REGION Network 151: PRODUCTION HOLD PB NOT RESET
   RUNG wire#powerrail
      Contact( "reset" )
      { S7_Templates := "SrcType := Word" } EQ_Contact(in1 := "DB101_DB_SDC_FAULTS".Carrier_Fault[44], in2 := 103)
      Coil( "DB302_HMI_Faults".Carrier44_Faults_3.%X14 )
   END_RUNG
   // the same network as SCL:
   "DB302_HMI_Faults".Carrier44_Faults_3.%X14 := "reset" AND ("DB101_DB_SDC_FAULTS".Carrier_Fault[44] = 103);
END_REGION

REGION Network 152: CARRIER FAULTS MASKED
   Label( C44_Comm_Flt )
   RUNG wire#powerrail
      Contact( "EMS".Carrier[44].FaultsMasked )
      Coil( "DB302_HMI_Faults".Carrier44_Faults_3.%X15 )
   END_RUNG
   // the same network as SCL:
   C44_Comm_Flt:
   "DB302_HMI_Faults".Carrier44_Faults_3.%X15 := "EMS".Carrier[44].FaultsMasked;
END_REGION

REGION Network 153: CARRIER 45 FAULTS
END_REGION

REGION Network 154: CARRIER PLC NOT COMMUNICATING
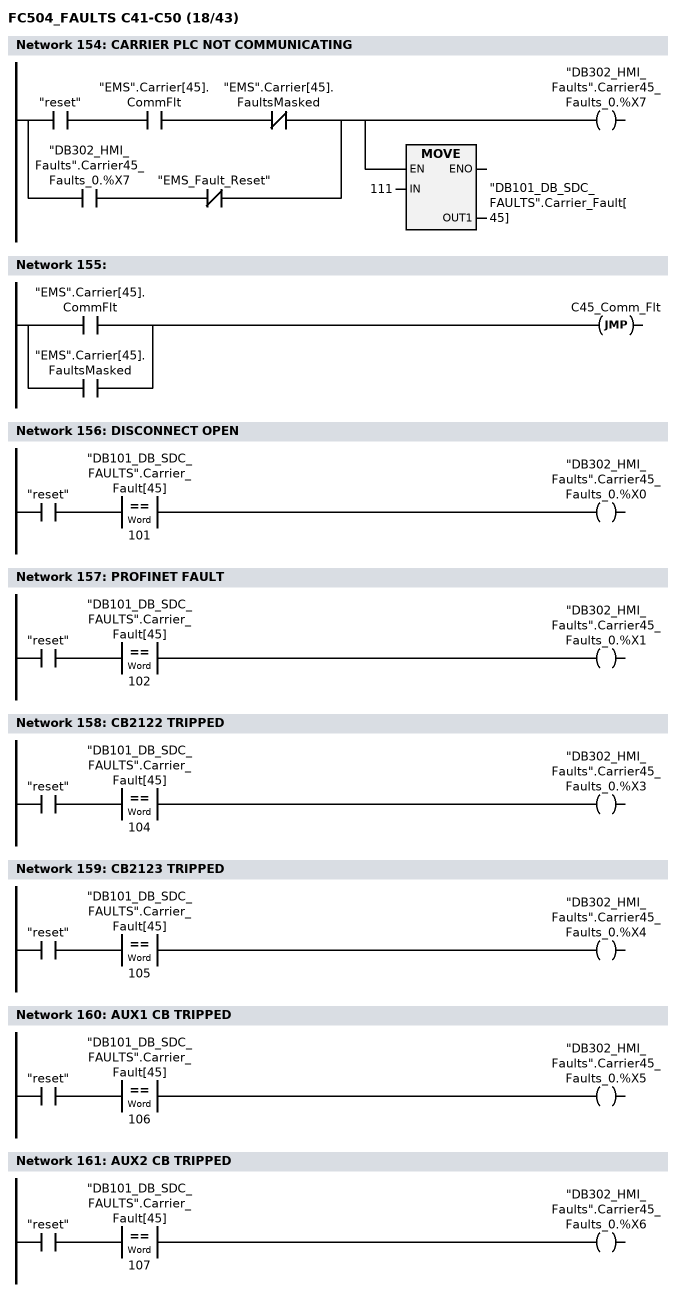
   RUNG wire#powerrail
      Contact( "reset" )
      Contact( "EMS".Carrier[45].CommFlt )
      I_Contact( "EMS".Carrier[45].FaultsMasked )
      wire#w1
      Coil( "DB302_HMI_Faults".Carrier45_Faults_0.%X7 )
   END_RUNG
   RUNG wire#powerrail
      Contact( "DB302_HMI_Faults".Carrier45_Faults_0.%X7 )
      I_Contact( "EMS_Fault_Reset" )
   END_RUNG wire#w1
   RUNG wire#w1
      Move(in := 111, out1 => "DB101_DB_SDC_FAULTS".Carrier_Fault[45])
   END_RUNG
   // the same network as SCL:
   "DB302_HMI_Faults".Carrier45_Faults_0.%X7 := ("reset" AND "EMS".Carrier[45].CommFlt AND NOT "EMS".Carrier[45].FaultsMasked) OR ("DB302_HMI_Faults".Carrier45_Faults_0.%X7 AND NOT "EMS_Fault_Reset");
   IF "DB302_HMI_Faults".Carrier45_Faults_0.%X7 THEN "DB101_DB_SDC_FAULTS".Carrier_Fault[45] := 111; END_IF;
END_REGION

REGION Network 155
   RUNG wire#powerrail
      Contact( "EMS".Carrier[45].CommFlt )
      wire#w1
      JumpCoil( C45_Comm_Flt )
   END_RUNG
   RUNG wire#powerrail
      Contact( "EMS".Carrier[45].FaultsMasked )
   END_RUNG wire#w1
   // the same network as SCL:
   IF "EMS".Carrier[45].CommFlt OR "EMS".Carrier[45].FaultsMasked THEN GOTO C45_Comm_Flt; END_IF;
END_REGION

REGION Network 156: DISCONNECT OPEN
   RUNG wire#powerrail
      Contact( "reset" )
      { S7_Templates := "SrcType := Word" } EQ_Contact(in1 := "DB101_DB_SDC_FAULTS".Carrier_Fault[45], in2 := 101)
      Coil( "DB302_HMI_Faults".Carrier45_Faults_0.%X0 )
   END_RUNG
   // the same network as SCL:
   "DB302_HMI_Faults".Carrier45_Faults_0.%X0 := "reset" AND ("DB101_DB_SDC_FAULTS".Carrier_Fault[45] = 101);
END_REGION

REGION Network 157: PROFINET FAULT
   RUNG wire#powerrail
      Contact( "reset" )
      { S7_Templates := "SrcType := Word" } EQ_Contact(in1 := "DB101_DB_SDC_FAULTS".Carrier_Fault[45], in2 := 102)
      Coil( "DB302_HMI_Faults".Carrier45_Faults_0.%X1 )
   END_RUNG
   // the same network as SCL:
   "DB302_HMI_Faults".Carrier45_Faults_0.%X1 := "reset" AND ("DB101_DB_SDC_FAULTS".Carrier_Fault[45] = 102);
END_REGION

REGION Network 158: CB2122 TRIPPED
   RUNG wire#powerrail
      Contact( "reset" )
      { S7_Templates := "SrcType := Word" } EQ_Contact(in1 := "DB101_DB_SDC_FAULTS".Carrier_Fault[45], in2 := 104)
      Coil( "DB302_HMI_Faults".Carrier45_Faults_0.%X3 )
   END_RUNG
   // the same network as SCL:
   "DB302_HMI_Faults".Carrier45_Faults_0.%X3 := "reset" AND ("DB101_DB_SDC_FAULTS".Carrier_Fault[45] = 104);
END_REGION

REGION Network 159: CB2123 TRIPPED
   RUNG wire#powerrail
      Contact( "reset" )
      { S7_Templates := "SrcType := Word" } EQ_Contact(in1 := "DB101_DB_SDC_FAULTS".Carrier_Fault[45], in2 := 105)
      Coil( "DB302_HMI_Faults".Carrier45_Faults_0.%X4 )
   END_RUNG
   // the same network as SCL:
   "DB302_HMI_Faults".Carrier45_Faults_0.%X4 := "reset" AND ("DB101_DB_SDC_FAULTS".Carrier_Fault[45] = 105);
END_REGION

REGION Network 160: AUX1 CB TRIPPED
   RUNG wire#powerrail
      Contact( "reset" )
      { S7_Templates := "SrcType := Word" } EQ_Contact(in1 := "DB101_DB_SDC_FAULTS".Carrier_Fault[45], in2 := 106)
      Coil( "DB302_HMI_Faults".Carrier45_Faults_0.%X5 )
   END_RUNG
   // the same network as SCL:
   "DB302_HMI_Faults".Carrier45_Faults_0.%X5 := "reset" AND ("DB101_DB_SDC_FAULTS".Carrier_Fault[45] = 106);
END_REGION

REGION Network 161: AUX2 CB TRIPPED
   RUNG wire#powerrail
      Contact( "reset" )
      { S7_Templates := "SrcType := Word" } EQ_Contact(in1 := "DB101_DB_SDC_FAULTS".Carrier_Fault[45], in2 := 107)
      Coil( "DB302_HMI_Faults".Carrier45_Faults_0.%X6 )
   END_RUNG
   // the same network as SCL:
   "DB302_HMI_Faults".Carrier45_Faults_0.%X6 := "reset" AND ("DB101_DB_SDC_FAULTS".Carrier_Fault[45] = 107);
END_REGION

REGION Network 162: SAFE INPUT CARD FAULT
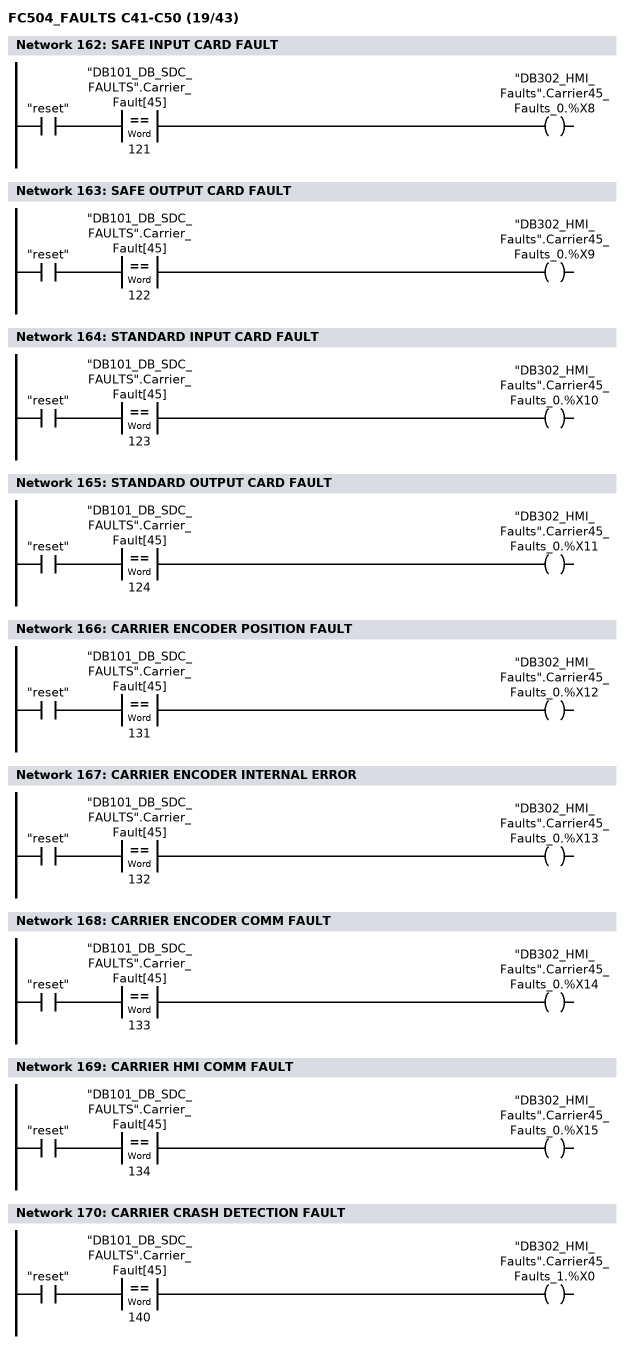
   RUNG wire#powerrail
      Contact( "reset" )
      { S7_Templates := "SrcType := Word" } EQ_Contact(in1 := "DB101_DB_SDC_FAULTS".Carrier_Fault[45], in2 := 121)
      Coil( "DB302_HMI_Faults".Carrier45_Faults_0.%X8 )
   END_RUNG
   // the same network as SCL:
   "DB302_HMI_Faults".Carrier45_Faults_0.%X8 := "reset" AND ("DB101_DB_SDC_FAULTS".Carrier_Fault[45] = 121);
END_REGION

REGION Network 163: SAFE OUTPUT CARD FAULT
   RUNG wire#powerrail
      Contact( "reset" )
      { S7_Templates := "SrcType := Word" } EQ_Contact(in1 := "DB101_DB_SDC_FAULTS".Carrier_Fault[45], in2 := 122)
      Coil( "DB302_HMI_Faults".Carrier45_Faults_0.%X9 )
   END_RUNG
   // the same network as SCL:
   "DB302_HMI_Faults".Carrier45_Faults_0.%X9 := "reset" AND ("DB101_DB_SDC_FAULTS".Carrier_Fault[45] = 122);
END_REGION

REGION Network 164: STANDARD INPUT CARD FAULT
   RUNG wire#powerrail
      Contact( "reset" )
      { S7_Templates := "SrcType := Word" } EQ_Contact(in1 := "DB101_DB_SDC_FAULTS".Carrier_Fault[45], in2 := 123)
      Coil( "DB302_HMI_Faults".Carrier45_Faults_0.%X10 )
   END_RUNG
   // the same network as SCL:
   "DB302_HMI_Faults".Carrier45_Faults_0.%X10 := "reset" AND ("DB101_DB_SDC_FAULTS".Carrier_Fault[45] = 123);
END_REGION

REGION Network 165: STANDARD OUTPUT CARD FAULT
   RUNG wire#powerrail
      Contact( "reset" )
      { S7_Templates := "SrcType := Word" } EQ_Contact(in1 := "DB101_DB_SDC_FAULTS".Carrier_Fault[45], in2 := 124)
      Coil( "DB302_HMI_Faults".Carrier45_Faults_0.%X11 )
   END_RUNG
   // the same network as SCL:
   "DB302_HMI_Faults".Carrier45_Faults_0.%X11 := "reset" AND ("DB101_DB_SDC_FAULTS".Carrier_Fault[45] = 124);
END_REGION

REGION Network 166: CARRIER ENCODER POSITION FAULT
   RUNG wire#powerrail
      Contact( "reset" )
      { S7_Templates := "SrcType := Word" } EQ_Contact(in1 := "DB101_DB_SDC_FAULTS".Carrier_Fault[45], in2 := 131)
      Coil( "DB302_HMI_Faults".Carrier45_Faults_0.%X12 )
   END_RUNG
   // the same network as SCL:
   "DB302_HMI_Faults".Carrier45_Faults_0.%X12 := "reset" AND ("DB101_DB_SDC_FAULTS".Carrier_Fault[45] = 131);
END_REGION

REGION Network 167: CARRIER ENCODER INTERNAL ERROR
   RUNG wire#powerrail
      Contact( "reset" )
      { S7_Templates := "SrcType := Word" } EQ_Contact(in1 := "DB101_DB_SDC_FAULTS".Carrier_Fault[45], in2 := 132)
      Coil( "DB302_HMI_Faults".Carrier45_Faults_0.%X13 )
   END_RUNG
   // the same network as SCL:
   "DB302_HMI_Faults".Carrier45_Faults_0.%X13 := "reset" AND ("DB101_DB_SDC_FAULTS".Carrier_Fault[45] = 132);
END_REGION

REGION Network 168: CARRIER ENCODER COMM FAULT
   RUNG wire#powerrail
      Contact( "reset" )
      { S7_Templates := "SrcType := Word" } EQ_Contact(in1 := "DB101_DB_SDC_FAULTS".Carrier_Fault[45], in2 := 133)
      Coil( "DB302_HMI_Faults".Carrier45_Faults_0.%X14 )
   END_RUNG
   // the same network as SCL:
   "DB302_HMI_Faults".Carrier45_Faults_0.%X14 := "reset" AND ("DB101_DB_SDC_FAULTS".Carrier_Fault[45] = 133);
END_REGION

REGION Network 169: CARRIER HMI COMM FAULT
   RUNG wire#powerrail
      Contact( "reset" )
      { S7_Templates := "SrcType := Word" } EQ_Contact(in1 := "DB101_DB_SDC_FAULTS".Carrier_Fault[45], in2 := 134)
      Coil( "DB302_HMI_Faults".Carrier45_Faults_0.%X15 )
   END_RUNG
   // the same network as SCL:
   "DB302_HMI_Faults".Carrier45_Faults_0.%X15 := "reset" AND ("DB101_DB_SDC_FAULTS".Carrier_Fault[45] = 134);
END_REGION

REGION Network 170: CARRIER CRASH DETECTION FAULT
   RUNG wire#powerrail
      Contact( "reset" )
      { S7_Templates := "SrcType := Word" } EQ_Contact(in1 := "DB101_DB_SDC_FAULTS".Carrier_Fault[45], in2 := 140)
      Coil( "DB302_HMI_Faults".Carrier45_Faults_1.%X0 )
   END_RUNG
   // the same network as SCL:
   "DB302_HMI_Faults".Carrier45_Faults_1.%X0 := "reset" AND ("DB101_DB_SDC_FAULTS".Carrier_Fault[45] = 140);
END_REGION

REGION Network 171: CARRIER NUMBER INVALID FAULT
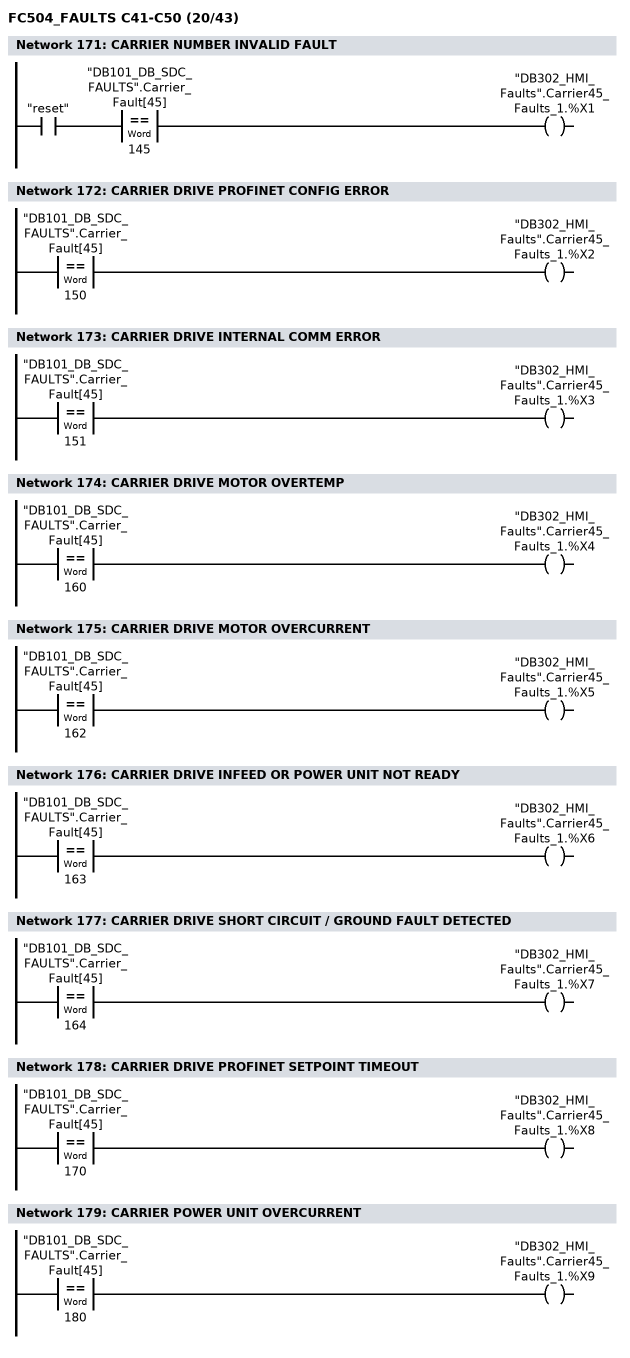
   RUNG wire#powerrail
      Contact( "reset" )
      { S7_Templates := "SrcType := Word" } EQ_Contact(in1 := "DB101_DB_SDC_FAULTS".Carrier_Fault[45], in2 := 145)
      Coil( "DB302_HMI_Faults".Carrier45_Faults_1.%X1 )
   END_RUNG
   // the same network as SCL:
   "DB302_HMI_Faults".Carrier45_Faults_1.%X1 := "reset" AND ("DB101_DB_SDC_FAULTS".Carrier_Fault[45] = 145);
END_REGION

REGION Network 172: CARRIER DRIVE PROFINET CONFIG ERROR
   RUNG wire#powerrail
      { S7_Templates := "SrcType := Word" } EQ_Contact(in1 := "DB101_DB_SDC_FAULTS".Carrier_Fault[45], in2 := 150)
      Coil( "DB302_HMI_Faults".Carrier45_Faults_1.%X2 )
   END_RUNG
   // the same network as SCL:
   "DB302_HMI_Faults".Carrier45_Faults_1.%X2 := "DB101_DB_SDC_FAULTS".Carrier_Fault[45] = 150;
END_REGION

REGION Network 173: CARRIER DRIVE INTERNAL COMM ERROR
   RUNG wire#powerrail
      { S7_Templates := "SrcType := Word" } EQ_Contact(in1 := "DB101_DB_SDC_FAULTS".Carrier_Fault[45], in2 := 151)
      Coil( "DB302_HMI_Faults".Carrier45_Faults_1.%X3 )
   END_RUNG
   // the same network as SCL:
   "DB302_HMI_Faults".Carrier45_Faults_1.%X3 := "DB101_DB_SDC_FAULTS".Carrier_Fault[45] = 151;
END_REGION

REGION Network 174: CARRIER DRIVE MOTOR OVERTEMP
   RUNG wire#powerrail
      { S7_Templates := "SrcType := Word" } EQ_Contact(in1 := "DB101_DB_SDC_FAULTS".Carrier_Fault[45], in2 := 160)
      Coil( "DB302_HMI_Faults".Carrier45_Faults_1.%X4 )
   END_RUNG
   // the same network as SCL:
   "DB302_HMI_Faults".Carrier45_Faults_1.%X4 := "DB101_DB_SDC_FAULTS".Carrier_Fault[45] = 160;
END_REGION

REGION Network 175: CARRIER DRIVE MOTOR OVERCURRENT
   RUNG wire#powerrail
      { S7_Templates := "SrcType := Word" } EQ_Contact(in1 := "DB101_DB_SDC_FAULTS".Carrier_Fault[45], in2 := 162)
      Coil( "DB302_HMI_Faults".Carrier45_Faults_1.%X5 )
   END_RUNG
   // the same network as SCL:
   "DB302_HMI_Faults".Carrier45_Faults_1.%X5 := "DB101_DB_SDC_FAULTS".Carrier_Fault[45] = 162;
END_REGION

REGION Network 176: CARRIER DRIVE INFEED OR POWER UNIT NOT READY
   RUNG wire#powerrail
      { S7_Templates := "SrcType := Word" } EQ_Contact(in1 := "DB101_DB_SDC_FAULTS".Carrier_Fault[45], in2 := 163)
      Coil( "DB302_HMI_Faults".Carrier45_Faults_1.%X6 )
   END_RUNG
   // the same network as SCL:
   "DB302_HMI_Faults".Carrier45_Faults_1.%X6 := "DB101_DB_SDC_FAULTS".Carrier_Fault[45] = 163;
END_REGION

REGION Network 177: CARRIER DRIVE SHORT CIRCUIT / GROUND FAULT DETECTED
   RUNG wire#powerrail
      { S7_Templates := "SrcType := Word" } EQ_Contact(in1 := "DB101_DB_SDC_FAULTS".Carrier_Fault[45], in2 := 164)
      Coil( "DB302_HMI_Faults".Carrier45_Faults_1.%X7 )
   END_RUNG
   // the same network as SCL:
   "DB302_HMI_Faults".Carrier45_Faults_1.%X7 := "DB101_DB_SDC_FAULTS".Carrier_Fault[45] = 164;
END_REGION

REGION Network 178: CARRIER DRIVE PROFINET SETPOINT TIMEOUT
   RUNG wire#powerrail
      { S7_Templates := "SrcType := Word" } EQ_Contact(in1 := "DB101_DB_SDC_FAULTS".Carrier_Fault[45], in2 := 170)
      Coil( "DB302_HMI_Faults".Carrier45_Faults_1.%X8 )
   END_RUNG
   // the same network as SCL:
   "DB302_HMI_Faults".Carrier45_Faults_1.%X8 := "DB101_DB_SDC_FAULTS".Carrier_Fault[45] = 170;
END_REGION

REGION Network 179: CARRIER POWER UNIT OVERCURRENT
   RUNG wire#powerrail
      { S7_Templates := "SrcType := Word" } EQ_Contact(in1 := "DB101_DB_SDC_FAULTS".Carrier_Fault[45], in2 := 180)
      Coil( "DB302_HMI_Faults".Carrier45_Faults_1.%X9 )
   END_RUNG
   // the same network as SCL:
   "DB302_HMI_Faults".Carrier45_Faults_1.%X9 := "DB101_DB_SDC_FAULTS".Carrier_Fault[45] = 180;
END_REGION

REGION Network 180: CARRIER POWER UNIT DC LINK OVERVOLTAGE
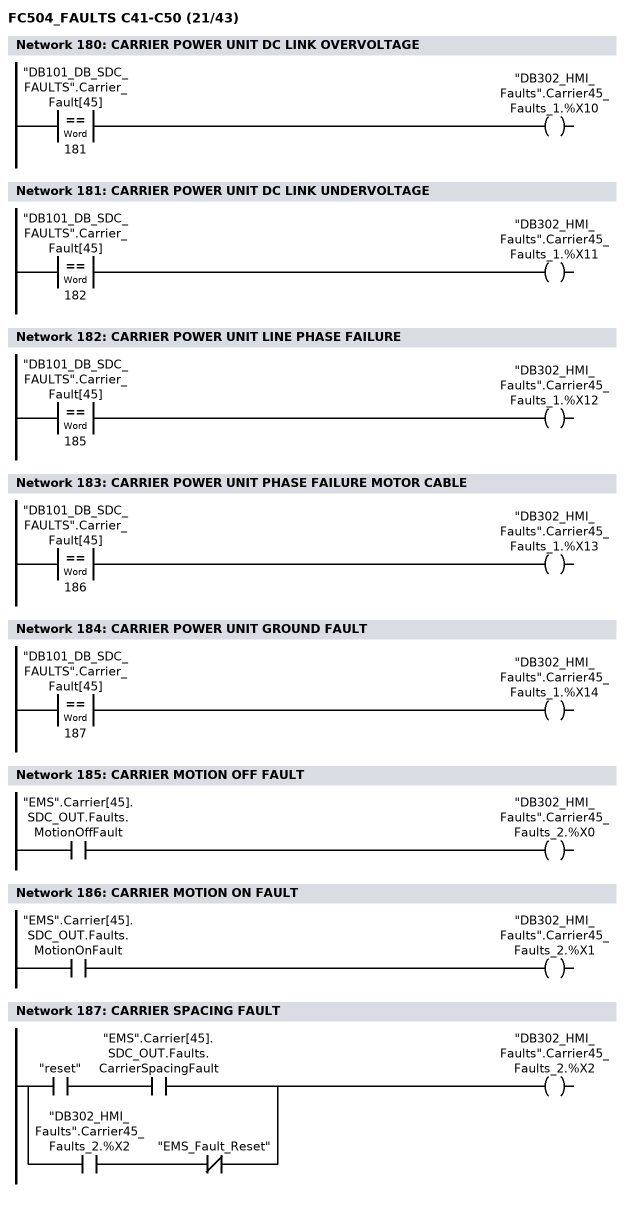
   RUNG wire#powerrail
      { S7_Templates := "SrcType := Word" } EQ_Contact(in1 := "DB101_DB_SDC_FAULTS".Carrier_Fault[45], in2 := 181)
      Coil( "DB302_HMI_Faults".Carrier45_Faults_1.%X10 )
   END_RUNG
   // the same network as SCL:
   "DB302_HMI_Faults".Carrier45_Faults_1.%X10 := "DB101_DB_SDC_FAULTS".Carrier_Fault[45] = 181;
END_REGION

REGION Network 181: CARRIER POWER UNIT DC LINK UNDERVOLTAGE
   RUNG wire#powerrail
      { S7_Templates := "SrcType := Word" } EQ_Contact(in1 := "DB101_DB_SDC_FAULTS".Carrier_Fault[45], in2 := 182)
      Coil( "DB302_HMI_Faults".Carrier45_Faults_1.%X11 )
   END_RUNG
   // the same network as SCL:
   "DB302_HMI_Faults".Carrier45_Faults_1.%X11 := "DB101_DB_SDC_FAULTS".Carrier_Fault[45] = 182;
END_REGION

REGION Network 182: CARRIER POWER UNIT LINE PHASE FAILURE
   RUNG wire#powerrail
      { S7_Templates := "SrcType := Word" } EQ_Contact(in1 := "DB101_DB_SDC_FAULTS".Carrier_Fault[45], in2 := 185)
      Coil( "DB302_HMI_Faults".Carrier45_Faults_1.%X12 )
   END_RUNG
   // the same network as SCL:
   "DB302_HMI_Faults".Carrier45_Faults_1.%X12 := "DB101_DB_SDC_FAULTS".Carrier_Fault[45] = 185;
END_REGION

REGION Network 183: CARRIER POWER UNIT PHASE FAILURE MOTOR CABLE
   RUNG wire#powerrail
      { S7_Templates := "SrcType := Word" } EQ_Contact(in1 := "DB101_DB_SDC_FAULTS".Carrier_Fault[45], in2 := 186)
      Coil( "DB302_HMI_Faults".Carrier45_Faults_1.%X13 )
   END_RUNG
   // the same network as SCL:
   "DB302_HMI_Faults".Carrier45_Faults_1.%X13 := "DB101_DB_SDC_FAULTS".Carrier_Fault[45] = 186;
END_REGION

REGION Network 184: CARRIER POWER UNIT GROUND FAULT
   RUNG wire#powerrail
      { S7_Templates := "SrcType := Word" } EQ_Contact(in1 := "DB101_DB_SDC_FAULTS".Carrier_Fault[45], in2 := 187)
      Coil( "DB302_HMI_Faults".Carrier45_Faults_1.%X14 )
   END_RUNG
   // the same network as SCL:
   "DB302_HMI_Faults".Carrier45_Faults_1.%X14 := "DB101_DB_SDC_FAULTS".Carrier_Fault[45] = 187;
END_REGION

REGION Network 185: CARRIER MOTION OFF FAULT
   RUNG wire#powerrail
      Contact( "EMS".Carrier[45].SDC_OUT.Faults.MotionOffFault )
      Coil( "DB302_HMI_Faults".Carrier45_Faults_2.%X0 )
   END_RUNG
   // the same network as SCL:
   "DB302_HMI_Faults".Carrier45_Faults_2.%X0 := "EMS".Carrier[45].SDC_OUT.Faults.MotionOffFault;
END_REGION

REGION Network 186: CARRIER MOTION ON FAULT
   RUNG wire#powerrail
      Contact( "EMS".Carrier[45].SDC_OUT.Faults.MotionOnFault )
      Coil( "DB302_HMI_Faults".Carrier45_Faults_2.%X1 )
   END_RUNG
   // the same network as SCL:
   "DB302_HMI_Faults".Carrier45_Faults_2.%X1 := "EMS".Carrier[45].SDC_OUT.Faults.MotionOnFault;
END_REGION

REGION Network 187: CARRIER SPACING FAULT
   RUNG wire#powerrail
      Contact( "reset" )
      Contact( "EMS".Carrier[45].SDC_OUT.Faults.CarrierSpacingFault )
      wire#w1
      Coil( "DB302_HMI_Faults".Carrier45_Faults_2.%X2 )
   END_RUNG
   RUNG wire#powerrail
      Contact( "DB302_HMI_Faults".Carrier45_Faults_2.%X2 )
      I_Contact( "EMS_Fault_Reset" )
   END_RUNG wire#w1
   // the same network as SCL:
   "DB302_HMI_Faults".Carrier45_Faults_2.%X2 := ("reset" AND "EMS".Carrier[45].SDC_OUT.Faults.CarrierSpacingFault) OR ("DB302_HMI_Faults".Carrier45_Faults_2.%X2 AND NOT "EMS_Fault_Reset");
END_REGION

REGION Network 188: DUPLICATE CARRIER NUMBER FAULT
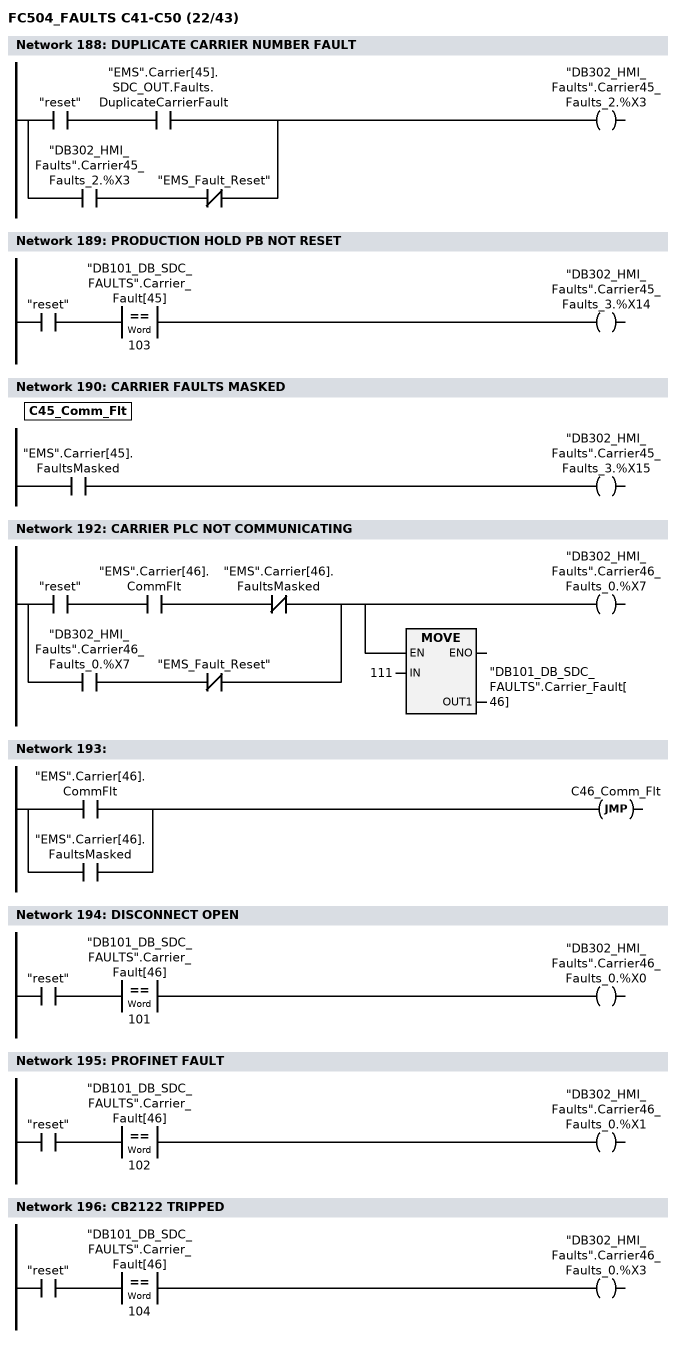
   RUNG wire#powerrail
      Contact( "reset" )
      Contact( "EMS".Carrier[45].SDC_OUT.Faults.DuplicateCarrierFault )
      wire#w1
      Coil( "DB302_HMI_Faults".Carrier45_Faults_2.%X3 )
   END_RUNG
   RUNG wire#powerrail
      Contact( "DB302_HMI_Faults".Carrier45_Faults_2.%X3 )
      I_Contact( "EMS_Fault_Reset" )
   END_RUNG wire#w1
   // the same network as SCL:
   "DB302_HMI_Faults".Carrier45_Faults_2.%X3 := ("reset" AND "EMS".Carrier[45].SDC_OUT.Faults.DuplicateCarrierFault) OR ("DB302_HMI_Faults".Carrier45_Faults_2.%X3 AND NOT "EMS_Fault_Reset");
END_REGION

REGION Network 189: PRODUCTION HOLD PB NOT RESET
   RUNG wire#powerrail
      Contact( "reset" )
      { S7_Templates := "SrcType := Word" } EQ_Contact(in1 := "DB101_DB_SDC_FAULTS".Carrier_Fault[45], in2 := 103)
      Coil( "DB302_HMI_Faults".Carrier45_Faults_3.%X14 )
   END_RUNG
   // the same network as SCL:
   "DB302_HMI_Faults".Carrier45_Faults_3.%X14 := "reset" AND ("DB101_DB_SDC_FAULTS".Carrier_Fault[45] = 103);
END_REGION

REGION Network 190: CARRIER FAULTS MASKED
   Label( C45_Comm_Flt )
   RUNG wire#powerrail
      Contact( "EMS".Carrier[45].FaultsMasked )
      Coil( "DB302_HMI_Faults".Carrier45_Faults_3.%X15 )
   END_RUNG
   // the same network as SCL:
   C45_Comm_Flt:
   "DB302_HMI_Faults".Carrier45_Faults_3.%X15 := "EMS".Carrier[45].FaultsMasked;
END_REGION

REGION Network 191: CARRIER 46 FAULTS
END_REGION

REGION Network 192: CARRIER PLC NOT COMMUNICATING
   RUNG wire#powerrail
      Contact( "reset" )
      Contact( "EMS".Carrier[46].CommFlt )
      I_Contact( "EMS".Carrier[46].FaultsMasked )
      wire#w1
      Coil( "DB302_HMI_Faults".Carrier46_Faults_0.%X7 )
   END_RUNG
   RUNG wire#powerrail
      Contact( "DB302_HMI_Faults".Carrier46_Faults_0.%X7 )
      I_Contact( "EMS_Fault_Reset" )
   END_RUNG wire#w1
   RUNG wire#w1
      Move(in := 111, out1 => "DB101_DB_SDC_FAULTS".Carrier_Fault[46])
   END_RUNG
   // the same network as SCL:
   "DB302_HMI_Faults".Carrier46_Faults_0.%X7 := ("reset" AND "EMS".Carrier[46].CommFlt AND NOT "EMS".Carrier[46].FaultsMasked) OR ("DB302_HMI_Faults".Carrier46_Faults_0.%X7 AND NOT "EMS_Fault_Reset");
   IF "DB302_HMI_Faults".Carrier46_Faults_0.%X7 THEN "DB101_DB_SDC_FAULTS".Carrier_Fault[46] := 111; END_IF;
END_REGION

REGION Network 193
   RUNG wire#powerrail
      Contact( "EMS".Carrier[46].CommFlt )
      wire#w1
      JumpCoil( C46_Comm_Flt )
   END_RUNG
   RUNG wire#powerrail
      Contact( "EMS".Carrier[46].FaultsMasked )
   END_RUNG wire#w1
   // the same network as SCL:
   IF "EMS".Carrier[46].CommFlt OR "EMS".Carrier[46].FaultsMasked THEN GOTO C46_Comm_Flt; END_IF;
END_REGION

REGION Network 194: DISCONNECT OPEN
   RUNG wire#powerrail
      Contact( "reset" )
      { S7_Templates := "SrcType := Word" } EQ_Contact(in1 := "DB101_DB_SDC_FAULTS".Carrier_Fault[46], in2 := 101)
      Coil( "DB302_HMI_Faults".Carrier46_Faults_0.%X0 )
   END_RUNG
   // the same network as SCL:
   "DB302_HMI_Faults".Carrier46_Faults_0.%X0 := "reset" AND ("DB101_DB_SDC_FAULTS".Carrier_Fault[46] = 101);
END_REGION

REGION Network 195: PROFINET FAULT
   RUNG wire#powerrail
      Contact( "reset" )
      { S7_Templates := "SrcType := Word" } EQ_Contact(in1 := "DB101_DB_SDC_FAULTS".Carrier_Fault[46], in2 := 102)
      Coil( "DB302_HMI_Faults".Carrier46_Faults_0.%X1 )
   END_RUNG
   // the same network as SCL:
   "DB302_HMI_Faults".Carrier46_Faults_0.%X1 := "reset" AND ("DB101_DB_SDC_FAULTS".Carrier_Fault[46] = 102);
END_REGION

REGION Network 196: CB2122 TRIPPED
   RUNG wire#powerrail
      Contact( "reset" )
      { S7_Templates := "SrcType := Word" } EQ_Contact(in1 := "DB101_DB_SDC_FAULTS".Carrier_Fault[46], in2 := 104)
      Coil( "DB302_HMI_Faults".Carrier46_Faults_0.%X3 )
   END_RUNG
   // the same network as SCL:
   "DB302_HMI_Faults".Carrier46_Faults_0.%X3 := "reset" AND ("DB101_DB_SDC_FAULTS".Carrier_Fault[46] = 104);
END_REGION

REGION Network 197: CB2123 TRIPPED
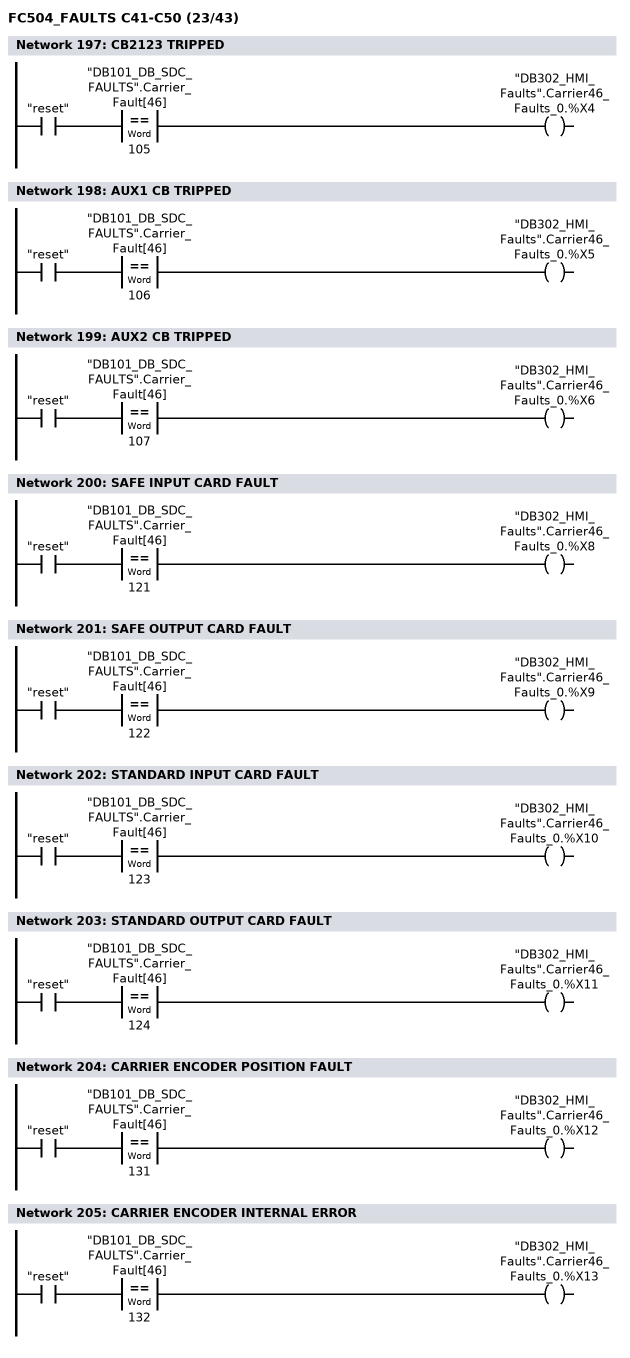
   RUNG wire#powerrail
      Contact( "reset" )
      { S7_Templates := "SrcType := Word" } EQ_Contact(in1 := "DB101_DB_SDC_FAULTS".Carrier_Fault[46], in2 := 105)
      Coil( "DB302_HMI_Faults".Carrier46_Faults_0.%X4 )
   END_RUNG
   // the same network as SCL:
   "DB302_HMI_Faults".Carrier46_Faults_0.%X4 := "reset" AND ("DB101_DB_SDC_FAULTS".Carrier_Fault[46] = 105);
END_REGION

REGION Network 198: AUX1 CB TRIPPED
   RUNG wire#powerrail
      Contact( "reset" )
      { S7_Templates := "SrcType := Word" } EQ_Contact(in1 := "DB101_DB_SDC_FAULTS".Carrier_Fault[46], in2 := 106)
      Coil( "DB302_HMI_Faults".Carrier46_Faults_0.%X5 )
   END_RUNG
   // the same network as SCL:
   "DB302_HMI_Faults".Carrier46_Faults_0.%X5 := "reset" AND ("DB101_DB_SDC_FAULTS".Carrier_Fault[46] = 106);
END_REGION

REGION Network 199: AUX2 CB TRIPPED
   RUNG wire#powerrail
      Contact( "reset" )
      { S7_Templates := "SrcType := Word" } EQ_Contact(in1 := "DB101_DB_SDC_FAULTS".Carrier_Fault[46], in2 := 107)
      Coil( "DB302_HMI_Faults".Carrier46_Faults_0.%X6 )
   END_RUNG
   // the same network as SCL:
   "DB302_HMI_Faults".Carrier46_Faults_0.%X6 := "reset" AND ("DB101_DB_SDC_FAULTS".Carrier_Fault[46] = 107);
END_REGION

REGION Network 200: SAFE INPUT CARD FAULT
   RUNG wire#powerrail
      Contact( "reset" )
      { S7_Templates := "SrcType := Word" } EQ_Contact(in1 := "DB101_DB_SDC_FAULTS".Carrier_Fault[46], in2 := 121)
      Coil( "DB302_HMI_Faults".Carrier46_Faults_0.%X8 )
   END_RUNG
   // the same network as SCL:
   "DB302_HMI_Faults".Carrier46_Faults_0.%X8 := "reset" AND ("DB101_DB_SDC_FAULTS".Carrier_Fault[46] = 121);
END_REGION

REGION Network 201: SAFE OUTPUT CARD FAULT
   RUNG wire#powerrail
      Contact( "reset" )
      { S7_Templates := "SrcType := Word" } EQ_Contact(in1 := "DB101_DB_SDC_FAULTS".Carrier_Fault[46], in2 := 122)
      Coil( "DB302_HMI_Faults".Carrier46_Faults_0.%X9 )
   END_RUNG
   // the same network as SCL:
   "DB302_HMI_Faults".Carrier46_Faults_0.%X9 := "reset" AND ("DB101_DB_SDC_FAULTS".Carrier_Fault[46] = 122);
END_REGION

REGION Network 202: STANDARD INPUT CARD FAULT
   RUNG wire#powerrail
      Contact( "reset" )
      { S7_Templates := "SrcType := Word" } EQ_Contact(in1 := "DB101_DB_SDC_FAULTS".Carrier_Fault[46], in2 := 123)
      Coil( "DB302_HMI_Faults".Carrier46_Faults_0.%X10 )
   END_RUNG
   // the same network as SCL:
   "DB302_HMI_Faults".Carrier46_Faults_0.%X10 := "reset" AND ("DB101_DB_SDC_FAULTS".Carrier_Fault[46] = 123);
END_REGION

REGION Network 203: STANDARD OUTPUT CARD FAULT
   RUNG wire#powerrail
      Contact( "reset" )
      { S7_Templates := "SrcType := Word" } EQ_Contact(in1 := "DB101_DB_SDC_FAULTS".Carrier_Fault[46], in2 := 124)
      Coil( "DB302_HMI_Faults".Carrier46_Faults_0.%X11 )
   END_RUNG
   // the same network as SCL:
   "DB302_HMI_Faults".Carrier46_Faults_0.%X11 := "reset" AND ("DB101_DB_SDC_FAULTS".Carrier_Fault[46] = 124);
END_REGION

REGION Network 204: CARRIER ENCODER POSITION FAULT
   RUNG wire#powerrail
      Contact( "reset" )
      { S7_Templates := "SrcType := Word" } EQ_Contact(in1 := "DB101_DB_SDC_FAULTS".Carrier_Fault[46], in2 := 131)
      Coil( "DB302_HMI_Faults".Carrier46_Faults_0.%X12 )
   END_RUNG
   // the same network as SCL:
   "DB302_HMI_Faults".Carrier46_Faults_0.%X12 := "reset" AND ("DB101_DB_SDC_FAULTS".Carrier_Fault[46] = 131);
END_REGION

REGION Network 205: CARRIER ENCODER INTERNAL ERROR
   RUNG wire#powerrail
      Contact( "reset" )
      { S7_Templates := "SrcType := Word" } EQ_Contact(in1 := "DB101_DB_SDC_FAULTS".Carrier_Fault[46], in2 := 132)
      Coil( "DB302_HMI_Faults".Carrier46_Faults_0.%X13 )
   END_RUNG
   // the same network as SCL:
   "DB302_HMI_Faults".Carrier46_Faults_0.%X13 := "reset" AND ("DB101_DB_SDC_FAULTS".Carrier_Fault[46] = 132);
END_REGION

REGION Network 206: CARRIER ENCODER COMM FAULT
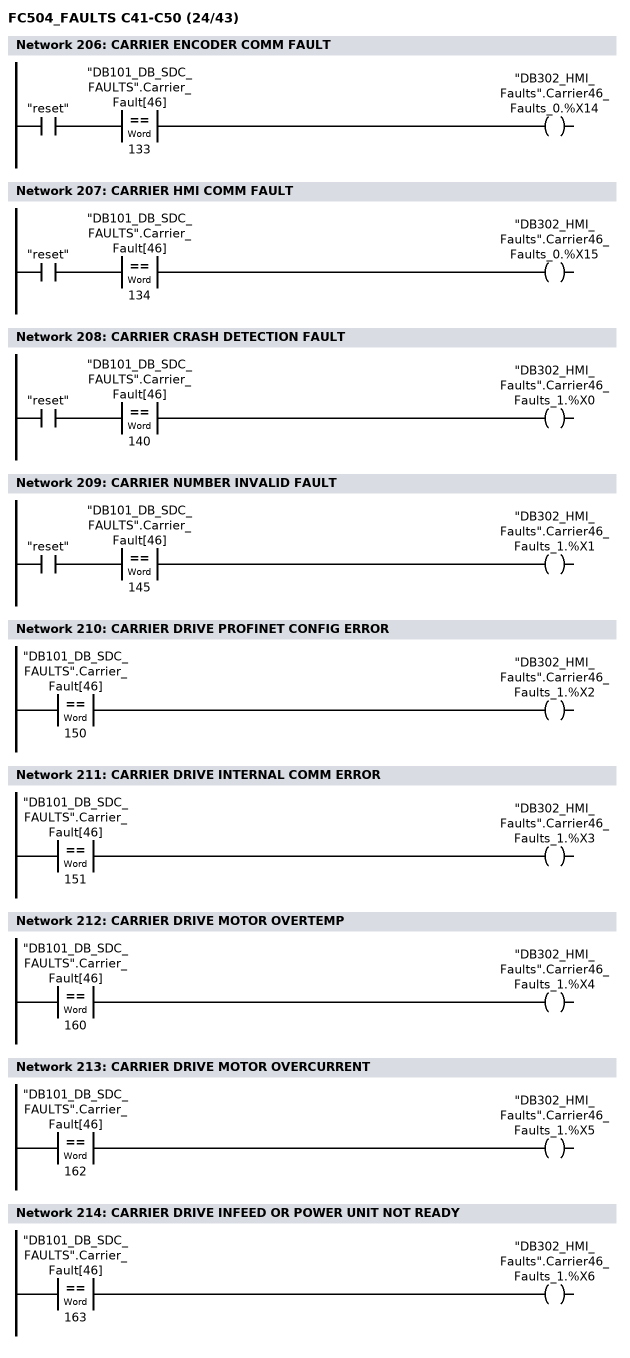
   RUNG wire#powerrail
      Contact( "reset" )
      { S7_Templates := "SrcType := Word" } EQ_Contact(in1 := "DB101_DB_SDC_FAULTS".Carrier_Fault[46], in2 := 133)
      Coil( "DB302_HMI_Faults".Carrier46_Faults_0.%X14 )
   END_RUNG
   // the same network as SCL:
   "DB302_HMI_Faults".Carrier46_Faults_0.%X14 := "reset" AND ("DB101_DB_SDC_FAULTS".Carrier_Fault[46] = 133);
END_REGION

REGION Network 207: CARRIER HMI COMM FAULT
   RUNG wire#powerrail
      Contact( "reset" )
      { S7_Templates := "SrcType := Word" } EQ_Contact(in1 := "DB101_DB_SDC_FAULTS".Carrier_Fault[46], in2 := 134)
      Coil( "DB302_HMI_Faults".Carrier46_Faults_0.%X15 )
   END_RUNG
   // the same network as SCL:
   "DB302_HMI_Faults".Carrier46_Faults_0.%X15 := "reset" AND ("DB101_DB_SDC_FAULTS".Carrier_Fault[46] = 134);
END_REGION

REGION Network 208: CARRIER CRASH DETECTION FAULT
   RUNG wire#powerrail
      Contact( "reset" )
      { S7_Templates := "SrcType := Word" } EQ_Contact(in1 := "DB101_DB_SDC_FAULTS".Carrier_Fault[46], in2 := 140)
      Coil( "DB302_HMI_Faults".Carrier46_Faults_1.%X0 )
   END_RUNG
   // the same network as SCL:
   "DB302_HMI_Faults".Carrier46_Faults_1.%X0 := "reset" AND ("DB101_DB_SDC_FAULTS".Carrier_Fault[46] = 140);
END_REGION

REGION Network 209: CARRIER NUMBER INVALID FAULT
   RUNG wire#powerrail
      Contact( "reset" )
      { S7_Templates := "SrcType := Word" } EQ_Contact(in1 := "DB101_DB_SDC_FAULTS".Carrier_Fault[46], in2 := 145)
      Coil( "DB302_HMI_Faults".Carrier46_Faults_1.%X1 )
   END_RUNG
   // the same network as SCL:
   "DB302_HMI_Faults".Carrier46_Faults_1.%X1 := "reset" AND ("DB101_DB_SDC_FAULTS".Carrier_Fault[46] = 145);
END_REGION

REGION Network 210: CARRIER DRIVE PROFINET CONFIG ERROR
   RUNG wire#powerrail
      { S7_Templates := "SrcType := Word" } EQ_Contact(in1 := "DB101_DB_SDC_FAULTS".Carrier_Fault[46], in2 := 150)
      Coil( "DB302_HMI_Faults".Carrier46_Faults_1.%X2 )
   END_RUNG
   // the same network as SCL:
   "DB302_HMI_Faults".Carrier46_Faults_1.%X2 := "DB101_DB_SDC_FAULTS".Carrier_Fault[46] = 150;
END_REGION

REGION Network 211: CARRIER DRIVE INTERNAL COMM ERROR
   RUNG wire#powerrail
      { S7_Templates := "SrcType := Word" } EQ_Contact(in1 := "DB101_DB_SDC_FAULTS".Carrier_Fault[46], in2 := 151)
      Coil( "DB302_HMI_Faults".Carrier46_Faults_1.%X3 )
   END_RUNG
   // the same network as SCL:
   "DB302_HMI_Faults".Carrier46_Faults_1.%X3 := "DB101_DB_SDC_FAULTS".Carrier_Fault[46] = 151;
END_REGION

REGION Network 212: CARRIER DRIVE MOTOR OVERTEMP
   RUNG wire#powerrail
      { S7_Templates := "SrcType := Word" } EQ_Contact(in1 := "DB101_DB_SDC_FAULTS".Carrier_Fault[46], in2 := 160)
      Coil( "DB302_HMI_Faults".Carrier46_Faults_1.%X4 )
   END_RUNG
   // the same network as SCL:
   "DB302_HMI_Faults".Carrier46_Faults_1.%X4 := "DB101_DB_SDC_FAULTS".Carrier_Fault[46] = 160;
END_REGION

REGION Network 213: CARRIER DRIVE MOTOR OVERCURRENT
   RUNG wire#powerrail
      { S7_Templates := "SrcType := Word" } EQ_Contact(in1 := "DB101_DB_SDC_FAULTS".Carrier_Fault[46], in2 := 162)
      Coil( "DB302_HMI_Faults".Carrier46_Faults_1.%X5 )
   END_RUNG
   // the same network as SCL:
   "DB302_HMI_Faults".Carrier46_Faults_1.%X5 := "DB101_DB_SDC_FAULTS".Carrier_Fault[46] = 162;
END_REGION

REGION Network 214: CARRIER DRIVE INFEED OR POWER UNIT NOT READY
   RUNG wire#powerrail
      { S7_Templates := "SrcType := Word" } EQ_Contact(in1 := "DB101_DB_SDC_FAULTS".Carrier_Fault[46], in2 := 163)
      Coil( "DB302_HMI_Faults".Carrier46_Faults_1.%X6 )
   END_RUNG
   // the same network as SCL:
   "DB302_HMI_Faults".Carrier46_Faults_1.%X6 := "DB101_DB_SDC_FAULTS".Carrier_Fault[46] = 163;
END_REGION

REGION Network 215: CARRIER DRIVE SHORT CIRCUIT / GROUND FAULT DETECTED
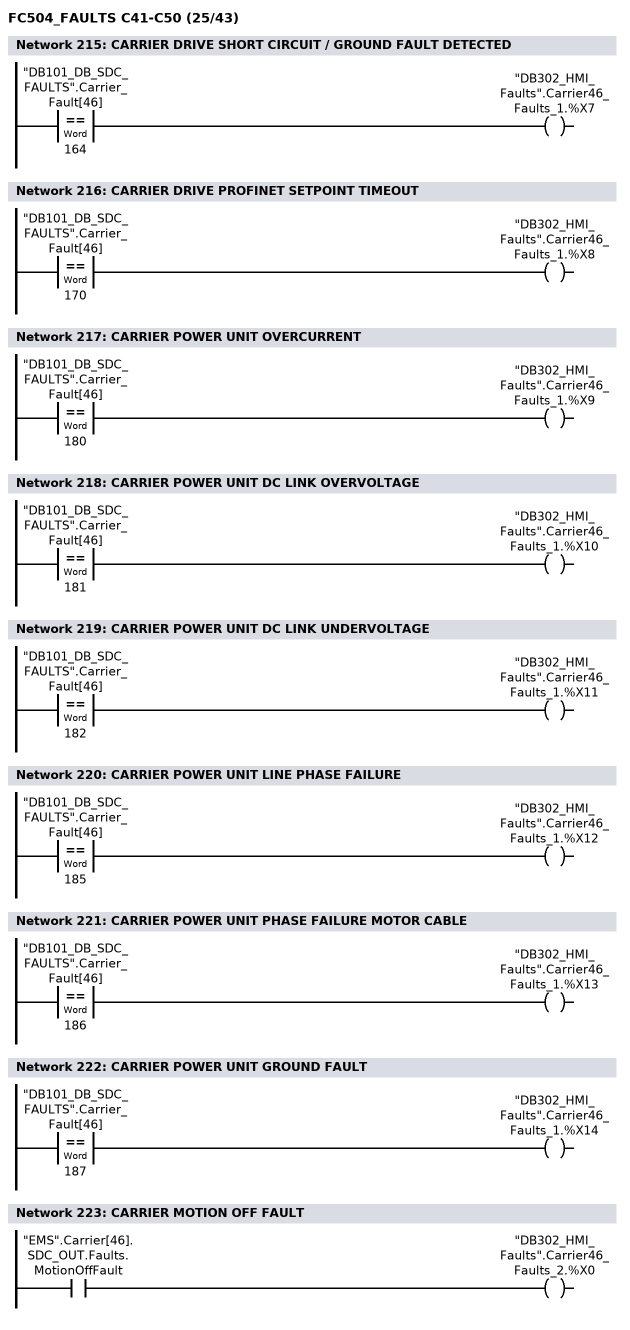
   RUNG wire#powerrail
      { S7_Templates := "SrcType := Word" } EQ_Contact(in1 := "DB101_DB_SDC_FAULTS".Carrier_Fault[46], in2 := 164)
      Coil( "DB302_HMI_Faults".Carrier46_Faults_1.%X7 )
   END_RUNG
   // the same network as SCL:
   "DB302_HMI_Faults".Carrier46_Faults_1.%X7 := "DB101_DB_SDC_FAULTS".Carrier_Fault[46] = 164;
END_REGION

REGION Network 216: CARRIER DRIVE PROFINET SETPOINT TIMEOUT
   RUNG wire#powerrail
      { S7_Templates := "SrcType := Word" } EQ_Contact(in1 := "DB101_DB_SDC_FAULTS".Carrier_Fault[46], in2 := 170)
      Coil( "DB302_HMI_Faults".Carrier46_Faults_1.%X8 )
   END_RUNG
   // the same network as SCL:
   "DB302_HMI_Faults".Carrier46_Faults_1.%X8 := "DB101_DB_SDC_FAULTS".Carrier_Fault[46] = 170;
END_REGION

REGION Network 217: CARRIER POWER UNIT OVERCURRENT
   RUNG wire#powerrail
      { S7_Templates := "SrcType := Word" } EQ_Contact(in1 := "DB101_DB_SDC_FAULTS".Carrier_Fault[46], in2 := 180)
      Coil( "DB302_HMI_Faults".Carrier46_Faults_1.%X9 )
   END_RUNG
   // the same network as SCL:
   "DB302_HMI_Faults".Carrier46_Faults_1.%X9 := "DB101_DB_SDC_FAULTS".Carrier_Fault[46] = 180;
END_REGION

REGION Network 218: CARRIER POWER UNIT DC LINK OVERVOLTAGE
   RUNG wire#powerrail
      { S7_Templates := "SrcType := Word" } EQ_Contact(in1 := "DB101_DB_SDC_FAULTS".Carrier_Fault[46], in2 := 181)
      Coil( "DB302_HMI_Faults".Carrier46_Faults_1.%X10 )
   END_RUNG
   // the same network as SCL:
   "DB302_HMI_Faults".Carrier46_Faults_1.%X10 := "DB101_DB_SDC_FAULTS".Carrier_Fault[46] = 181;
END_REGION

REGION Network 219: CARRIER POWER UNIT DC LINK UNDERVOLTAGE
   RUNG wire#powerrail
      { S7_Templates := "SrcType := Word" } EQ_Contact(in1 := "DB101_DB_SDC_FAULTS".Carrier_Fault[46], in2 := 182)
      Coil( "DB302_HMI_Faults".Carrier46_Faults_1.%X11 )
   END_RUNG
   // the same network as SCL:
   "DB302_HMI_Faults".Carrier46_Faults_1.%X11 := "DB101_DB_SDC_FAULTS".Carrier_Fault[46] = 182;
END_REGION

REGION Network 220: CARRIER POWER UNIT LINE PHASE FAILURE
   RUNG wire#powerrail
      { S7_Templates := "SrcType := Word" } EQ_Contact(in1 := "DB101_DB_SDC_FAULTS".Carrier_Fault[46], in2 := 185)
      Coil( "DB302_HMI_Faults".Carrier46_Faults_1.%X12 )
   END_RUNG
   // the same network as SCL:
   "DB302_HMI_Faults".Carrier46_Faults_1.%X12 := "DB101_DB_SDC_FAULTS".Carrier_Fault[46] = 185;
END_REGION

REGION Network 221: CARRIER POWER UNIT PHASE FAILURE MOTOR CABLE
   RUNG wire#powerrail
      { S7_Templates := "SrcType := Word" } EQ_Contact(in1 := "DB101_DB_SDC_FAULTS".Carrier_Fault[46], in2 := 186)
      Coil( "DB302_HMI_Faults".Carrier46_Faults_1.%X13 )
   END_RUNG
   // the same network as SCL:
   "DB302_HMI_Faults".Carrier46_Faults_1.%X13 := "DB101_DB_SDC_FAULTS".Carrier_Fault[46] = 186;
END_REGION

REGION Network 222: CARRIER POWER UNIT GROUND FAULT
   RUNG wire#powerrail
      { S7_Templates := "SrcType := Word" } EQ_Contact(in1 := "DB101_DB_SDC_FAULTS".Carrier_Fault[46], in2 := 187)
      Coil( "DB302_HMI_Faults".Carrier46_Faults_1.%X14 )
   END_RUNG
   // the same network as SCL:
   "DB302_HMI_Faults".Carrier46_Faults_1.%X14 := "DB101_DB_SDC_FAULTS".Carrier_Fault[46] = 187;
END_REGION

REGION Network 223: CARRIER MOTION OFF FAULT
   RUNG wire#powerrail
      Contact( "EMS".Carrier[46].SDC_OUT.Faults.MotionOffFault )
      Coil( "DB302_HMI_Faults".Carrier46_Faults_2.%X0 )
   END_RUNG
   // the same network as SCL:
   "DB302_HMI_Faults".Carrier46_Faults_2.%X0 := "EMS".Carrier[46].SDC_OUT.Faults.MotionOffFault;
END_REGION

REGION Network 224: CARRIER MOTION ON FAULT
